   "Carrier_17_SpareSafetyInput(2_4)" AT %I1214.4 : Bool;   // SPARE SAFETY INPUT
   "Carrier_17_SpareSafetyInput(2_5)" AT %I1214.5 : Bool;   // SPARE SAFETY INPUT
   "Carrier_17_SpareSafetyInput(2_6)" AT %I1214.6 : Bool;   // SPARE SAFETY INPUT
   "Carrier_17_SpareSafetyInput(2_7)" AT %I1214.7 : Bool;   // SPARE SAFETY INPUT
   "Carrier_17_Slot3_SafetyOutput" AT %IW1215 : Word;   // SLOT 3 SAFETY OUTPUT WORD
   "Carrier_17_Crash_Detect_OK" AT %I1215.0 : Bool;   // CARRIER CRASH DETECT
   "Carrier_17_SpareSafetyOutput(3_1)" AT %I1215.1 : Bool;   // SPARE SAFETY OUTPUT
   "Carrier_17_SpareSafetyOutput(3_2)" AT %I1215.2 : Bool;   // SPARE SAFETY OUTPUT
   "Carrier_17_SpareSafetyOutput(3_3)" AT %I1215.3 : Bool;   // SPARE SAFETY OUTPUT
   "Carrier_17_SpareSafetyOutput(3_4)" AT %I1215.4 : Bool;   // SPARE SAFETY OUTPUT
   "Carrier_17_SpareSafetyOutput(3_5)" AT %I1215.5 : Bool;   // SPARE SAFETY OUTPUT
   "Carrier_17_SpareSafetyOutput(3_6)" AT %I1215.6 : Bool;   // SPARE SAFETY OUTPUT
   "Carrier_17_SpareSafetyOutput(3_7)" AT %I1215.7 : Bool;   // SPARE SAFETY OUTPUT
   "Carrier_17_Slot4_Input" AT %IW1216 : Word;   // SLOT 4 INPUT WORD
   "Carrier_17_480VPowerOn_MDCB1" AT %I1216.0 : Bool;   // 480 VAC POWER ON MDCB 1
   "Carrier_17_SpareInput(4_1)" AT %I1216.1 : Bool;   // SPARE INPUT
   "Carrier_17_SpareInput(4_2)" AT %I1216.2 : Bool;   // SPARE INPUT
   "Carrier_17_SitopSelectStatus" AT %I1216.3 : Bool;   // SITOP SELECT STATUS
   "Carrier_17_DCsupplyOnPSCB2" AT %I1216.4 : Bool;   // DC SUPPLY ON PSCB 2
   "Carrier_17_SpareInput(4_5)" AT %I1216.5 : Bool;   // SPARE INPUT
   "Carrier_17_SpareInput(4_6)" AT %I1216.6 : Bool;   // SPARE INPUT
   "Carrier_17_SpareInput(4_7)" AT %I1216.7 : Bool;   // SPARE INPUT
   "Carrier_17_PB1_ProdHoldLH" AT %I1217.0 : Bool;   // PB 1 PRODUCTION HOLD LH
   "Carrier_17_PB2_ResetLH" AT %I1217.1 : Bool;   // PB 2 RESET LH
   "Carrier_17_PB3_ProdHoldRH" AT %I1217.2 : Bool;   // PB 3 PRODUCTION HOLD RH
   "Carrier_17_PB4_ResetRH" AT %I1217.3 : Bool;   // PB 4 RESET RH
   "Carrier_17_SpareInput(4_14)" AT %I1217.4 : Bool;   // SPARE INPUT
   "Carrier_17_SpareInput(4_15)" AT %I1217.5 : Bool;   // SPARE INPUT
   "Carrier_17_SpareInput(4_16)" AT %I1217.6 : Bool;   // SPARE INPUT
   "Carrier_17_SpareInput(4_17)" AT %I1217.7 : Bool;   // SPARE INPUT
   "Carrier_17_Slot5_Output" AT %IW1218 : Word;   // SLOT 5 OUTPUT WORD
   "Carrier_17_IRD400_HMI_24VDC_ENABLE" AT %I1218.0 : Bool;   // IRD 400 PANEL HMI 24V DC POWER
   "Carrier_17_FaultLight_LH" AT %I1218.1 : Bool;   // FAULT LIGHT LH
   "Carrier_17_RunLight_LH" AT %I1218.2 : Bool;   // RUN LIGHT LH
   "Carrier_17_FaultLight_RH" AT %I1218.3 : Bool;   // FAULT LIGHT RH
   "Carrier_17_RunLight_RH" AT %I1218.4 : Bool;   // RUN LIGHT RH
   "Carrier_17_SpareOutput(5_5)" AT %I1218.5 : Bool;   // SPARE OUTPUT
   "Carrier_17_SpareOutput(5_6)" AT %I1218.6 : Bool;   // SPARE OUTPUT
   "Carrier_17_SpareOutput(5_7)" AT %I1218.7 : Bool;   // SPARE OUTPUT
   "Carrier_17_ActualSpeed" AT %IW1220 : Word;   // ACTUAL SPEED
   "Carrier_17_CarrierDriveAlarm" AT %IW1222 : Word;   // CARRIER DRIVE ALARM
   "Carrier_17_CarrierDriveWarning" AT %IW1224 : Word;   // CARRIER DRIVE WARNING
   "Carrier_18_Status" AT %IW1250 : Word;   // CARRIER STATUS WORD
   "Carrier_18_Status.0" AT %I1250.0 : Bool;   // HEARTBEAT
   "Carrier_18_Status.1" AT %I1250.1 : Bool;   // MANUAL
   "Carrier_18_Status.2" AT %I1250.2 : Bool;   // IN_AUTO
   "Carrier_18_Status.3" AT %I1250.3 : Bool;   // POSITIONING_COMPLETE
   "Carrier_18_Status.4" AT %I1250.4 : Bool;   // PRODUCTION HOLD
   "Carrier_18_Status.5" AT %I1250.5 : Bool;   // CARRIER MOVING FORWARD
   "Carrier_18_Status.6" AT %I1250.6 : Bool;   // CARRIER MOVING REVERSE
   "Carrier_18_Status.7" AT %I1250.7 : Bool;   // CARRIER FAULT
   "Carrier_18_Status.8" AT %I1251.0 : Bool;   // CRASH DETECT TRIPPED
   "Carrier_18_Status.9" AT %I1251.1 : Bool;
   "Carrier_18_Status.10" AT %I1251.2 : Bool;
   "Carrier_18_Status.11" AT %I1251.3 : Bool;
   "Carrier_18_Status.12" AT %I1251.4 : Bool;
   "Carrier_18_Status.13" AT %I1251.5 : Bool;
   "Carrier_18_Status.14" AT %I1251.6 : Bool;
   "Carrier_18_Status.15" AT %I1251.7 : Bool;
   "Carrier_18_SDCFaultCode" AT %IW1252 : Word;   // SDC FAULT CODE
   "Carrier_18_CarrierPosition" AT %ID1254 : DWord;   // CARRIER POSITION
   "Carrier_18_CarrierNumber" AT %IW1258 : Word;   // CARRIER NUMBER
   "Carrier_18_G120DControlWord" AT %IW1260 : Word;   // G120D_STW1_CONTROL
   "Carrier_18_G120DControlWord.0" AT %I1260.0 : Bool;   // Bit_00_ON
   "Carrier_18_G120DControlWord.1" AT %I1260.1 : Bool;   // Bit_01_AUS2_INH
   "Carrier_18_G120DControlWord.2" AT %I1260.2 : Bool;   // Bit_02_AUS3_STOP
   "Carrier_18_G120DControlWord.3" AT %I1260.3 : Bool;   // Bit_03_EN
   "Carrier_18_G120DControlWord.4" AT %I1260.4 : Bool;   // Bit_04_EN_RAMP
   "Carrier_18_G120DControlWord.5" AT %I1260.5 : Bool;   // Bit_05_START_RAMP
   "Carrier_18_G120DControlWord.6" AT %I1260.6 : Bool;   // Bit_06_SETPOINT
   "Carrier_18_G120DControlWord.7" AT %I1260.7 : Bool;   // Bit_07_RESET
   "Carrier_18_G120DControlWord.8" AT %I1261.0 : Bool;   // Bit_08_JOG_R
   "Carrier_18_G120DControlWord.9" AT %I1261.1 : Bool;   // Bit_09_JOG_L
   "Carrier_18_G120DControlWord.10" AT %I1261.2 : Bool;   // Bit_10_CONTR_PLC
   "Carrier_18_G120DControlWord.11" AT %I1261.3 : Bool;   // Bit_11_REVERSE
   "Carrier_18_G120DControlWord.12" AT %I1261.4 : Bool;   // Bit_12_BRAKE_RELEASE
   "Carrier_18_G120DControlWord.13" AT %I1261.5 : Bool;   // Bit_13_DDS
   "Carrier_18_G120DControlWord.14" AT %I1261.6 : Bool;   // Bit_14_DO0
   "Carrier_18_G120DControlWord.15" AT %I1261.7 : Bool;   // Bit_15_DO1
   "Carrier_18_G120DStatusWord" AT %IW1262 : Word;   // G120D_ZSW1_STATUS
   "Carrier_18_G120DStatusWord.0" AT %I1262.0 : Bool;   // Bit_00_READY_RUN
   "Carrier_18_G120DStatusWord.1" AT %I1262.1 : Bool;   // Bit_01_READY_ON
   "Carrier_18_G120DStatusWord.2" AT %I1262.2 : Bool;   // Bit_02_ENABLE
   "Carrier_18_G120DStatusWord.3" AT %I1262.3 : Bool;   // Bit_03_FAULT
   "Carrier_18_G120DStatusWord.4" AT %I1262.4 : Bool;   // Bit_04_OFF2
   "Carrier_18_G120DStatusWord.5" AT %I1262.5 : Bool;   // Bit_05_OFF3
   "Carrier_18_G120DStatusWord.6" AT %I1262.6 : Bool;   // Bit_06_LOCK_OUT
   "Carrier_18_G120DStatusWord.7" AT %I1262.7 : Bool;   // Bit_07_WARN
   "Carrier_18_G120DStatusWord.8" AT %I1263.0 : Bool;   // Bit_08_NO_DEVIATION
   "Carrier_18_G120DStatusWord.9" AT %I1263.1 : Bool;   // Bit_09_CONTR_PLC
   "Carrier_18_G120DStatusWord.10" AT %I1263.2 : Bool;   // Bit_10_F_MAX
   "Carrier_18_G120DStatusWord.11" AT %I1263.3 : Bool;   // Bit_11_LIMIT_REACHED
   "Carrier_18_G120DStatusWord.12" AT %I1263.4 : Bool;   // Bit_12_BRAKE_OPEN
   "Carrier_18_G120DStatusWord.13" AT %I1263.5 : Bool;   // Bit_13_NO_OVERTEMP
   "Carrier_18_G120DStatusWord.14" AT %I1263.6 : Bool;   // Bit_14_CW_CCW
   "Carrier_18_G120DStatusWord.15" AT %I1263.7 : Bool;   // Bit_15_OVERL
   "Carrier_18_Slot2_Input" AT %IW1264 : Word;   // SLOT 2 INPUT WORD
   "Carrier_18_CrashDetectSW" AT %I1264.0 : Bool;   // CRASH DETECT SW
   "Carrier_18_SpareSafetyInput(2_1)" AT %I1264.1 : Bool;   // SPARE SAFETY INPUT
   "Carrier_18_SpareSafetyInput(2_2)" AT %I1264.2 : Bool;   // SPARE SAFETY INPUT
   "Carrier_18_SpareSafetyInput(2_3)" AT %I1264.3 : Bool;   // SPARE SAFETY INPUT
   "Carrier_18_SpareSafetyInput(2_4)" AT %I1264.4 : Bool;   // SPARE SAFETY INPUT
   "Carrier_18_SpareSafetyInput(2_5)" AT %I1264.5 : Bool;   // SPARE SAFETY INPUT
   "Carrier_18_SpareSafetyInput(2_6)" AT %I1264.6 : Bool;   // SPARE SAFETY INPUT
   "Carrier_18_SpareSafetyInput(2_7)" AT %I1264.7 : Bool;   // SPARE SAFETY INPUT
   "Carrier_18_Slot3_SafetyOutput" AT %IW1265 : Word;   // SLOT 3 SAFETY OUTPUT WORD
   "Carrier_18_Crash_Detect_OK" AT %I1265.0 : Bool;   // CARRIER CRASH DETECT
   "Carrier_18_SpareSafetyOutput(3_1)" AT %I1265.1 : Bool;   // SPARE SAFETY OUTPUT
   "Carrier_18_SpareSafetyOutput(3_2)" AT %I1265.2 : Bool;   // SPARE SAFETY OUTPUT
   "Carrier_18_SpareSafetyOutput(3_3)" AT %I1265.3 : Bool;   // SPARE SAFETY OUTPUT
   "Carrier_18_SpareSafetyOutput(3_4)" AT %I1265.4 : Bool;   // SPARE SAFETY OUTPUT
   "Carrier_18_SpareSafetyOutput(3_5)" AT %I1265.5 : Bool;   // SPARE SAFETY OUTPUT
   "Carrier_18_SpareSafetyOutput(3_6)" AT %I1265.6 : Bool;   // SPARE SAFETY OUTPUT
   "Carrier_18_SpareSafetyOutput(3_7)" AT %I1265.7 : Bool;   // SPARE SAFETY OUTPUT
   "Carrier_18_Slot4_Input" AT %IW1266 : Word;   // SLOT 4 INPUT WORD
   "Carrier_18_480VPowerOn_MDCB1" AT %I1266.0 : Bool;   // 480 VAC POWER ON MDCB 1
   "Carrier_18_SpareInput(4_1)" AT %I1266.1 : Bool;   // SPARE INPUT
   "Carrier_18_SpareInput(4_2)" AT %I1266.2 : Bool;   // SPARE INPUT
   "Carrier_18_SitopSelectStatus" AT %I1266.3 : Bool;   // SITOP SELECT STATUS
   "Carrier_18_DCsupplyOnPSCB2" AT %I1266.4 : Bool;   // DC SUPPLY ON PSCB 2
   "Carrier_18_SpareInput(4_5)" AT %I1266.5 : Bool;   // SPARE INPUT
   "Carrier_18_SpareInput(4_6)" AT %I1266.6 : Bool;   // SPARE INPUT
   "Carrier_18_SpareInput(4_7)" AT %I1266.7 : Bool;   // SPARE INPUT
   "Carrier_18_PB1_ProdHoldLH" AT %I1267.0 : Bool;   // PB 1 PRODUCTION HOLD LH
   "Carrier_18_PB2_ResetLH" AT %I1267.1 : Bool;   // PB 2 RESET LH
   "Carrier_18_PB3_ProdHoldRH" AT %I1267.2 : Bool;   // PB 3 PRODUCTION HOLD RH
   "Carrier_18_PB4_ResetRH" AT %I1267.3 : Bool;   // PB 4 RESET RH
   "Carrier_18_SpareInput(4_14)" AT %I1267.4 : Bool;   // SPARE INPUT
   "Carrier_18_SpareInput(4_15)" AT %I1267.5 : Bool;   // SPARE INPUT
   "Carrier_18_SpareInput(4_16)" AT %I1267.6 : Bool;   // SPARE INPUT
   "Carrier_18_SpareInput(4_17)" AT %I1267.7 : Bool;   // SPARE INPUT
   "Carrier_18_Slot5_Output" AT %IW1268 : Word;   // SLOT 5 OUTPUT WORD
   "Carrier_18_IRD400_HMI_24VDC_ENABLE" AT %I1268.0 : Bool;   // IRD 400 PANEL HMI 24V DC POWER
   "Carrier_18_FaultLight_LH" AT %I1268.1 : Bool;   // FAULT LIGHT LH
   "Carrier_18_RunLight_LH" AT %I1268.2 : Bool;   // RUN LIGHT LH
   "Carrier_18_FaultLight_RH" AT %I1268.3 : Bool;   // FAULT LIGHT RH
   "Carrier_18_RunLight_RH" AT %I1268.4 : Bool;   // RUN LIGHT RH
   "Carrier_18_SpareOutput(5_5)" AT %I1268.5 : Bool;   // SPARE OUTPUT
   "Carrier_18_SpareOutput(5_6)" AT %I1268.6 : Bool;   // SPARE OUTPUT
   "Carrier_18_SpareOutput(5_7)" AT %I1268.7 : Bool;   // SPARE OUTPUT
   "Carrier_18_ActualSpeed" AT %IW1270 : Word;   // ACTUAL SPEED
   "Carrier_18_CarrierDriveAlarm" AT %IW1272 : Word;   // CARRIER DRIVE ALARM
   "Carrier_18_CarrierDriveWarning" AT %IW1274 : Word;   // CARRIER DRIVE WARNING
   "Carrier_19_Status" AT %IW1300 : Word;   // CARRIER STATUS WORD
   "Carrier_19_Status.0" AT %I1300.0 : Bool;   // HEARTBEAT
   "Carrier_19_Status.1" AT %I1300.1 : Bool;   // MANUAL
   "Carrier_19_Status.2" AT %I1300.2 : Bool;   // IN_AUTO
   "Carrier_19_Status.3" AT %I1300.3 : Bool;   // POSITIONING_COMPLETE
   "Carrier_19_Status.4" AT %I1300.4 : Bool;   // PRODUCTION HOLD
   "Carrier_19_Status.5" AT %I1300.5 : Bool;   // CARRIER MOVING FORWARD
   "Carrier_19_Status.6" AT %I1300.6 : Bool;   // CARRIER MOVING REVERSE
   "Carrier_19_Status.7" AT %I1300.7 : Bool;   // CARRIER FAULT
   "Carrier_19_Status.8" AT %I1301.0 : Bool;   // CRASH DETECT TRIPPED
   "Carrier_19_Status.9" AT %I1301.1 : Bool;
   "Carrier_19_Status.10" AT %I1301.2 : Bool;
   "Carrier_19_Status.11" AT %I1301.3 : Bool;
   "Carrier_19_Status.12" AT %I1301.4 : Bool;
   "Carrier_19_Status.13" AT %I1301.5 : Bool;
   "Carrier_19_Status.14" AT %I1301.6 : Bool;
   "Carrier_19_Status.15" AT %I1301.7 : Bool;
   "Carrier_19_SDCFaultCode" AT %IW1302 : Word;   // SDC FAULT CODE
   "Carrier_19_CarrierPosition" AT %ID1304 : DWord;   // CARRIER POSITION
   "Carrier_19_CarrierNumber" AT %IW1308 : Word;   // CARRIER NUMBER
   "Carrier_19_G120DControlWord" AT %IW1310 : Word;   // G120D_STW1_CONTROL
   "Carrier_19_G120DControlWord.0" AT %I1310.0 : Bool;   // Bit_00_ON
   "Carrier_19_G120DControlWord.1" AT %I1310.1 : Bool;   // Bit_01_AUS2_INH
   "Carrier_19_G120DControlWord.2" AT %I1310.2 : Bool;   // Bit_02_AUS3_STOP
   "Carrier_19_G120DControlWord.3" AT %I1310.3 : Bool;   // Bit_03_EN
   "Carrier_19_G120DControlWord.4" AT %I1310.4 : Bool;   // Bit_04_EN_RAMP
   "Carrier_19_G120DControlWord.5" AT %I1310.5 : Bool;   // Bit_05_START_RAMP
   "Carrier_19_G120DControlWord.6" AT %I1310.6 : Bool;   // Bit_06_SETPOINT
   "Carrier_19_G120DControlWord.7" AT %I1310.7 : Bool;   // Bit_07_RESET
   "Carrier_19_G120DControlWord.8" AT %I1311.0 : Bool;   // Bit_08_JOG_R
   "Carrier_19_G120DControlWord.9" AT %I1311.1 : Bool;   // Bit_09_JOG_L
   "Carrier_19_G120DControlWord.10" AT %I1311.2 : Bool;   // Bit_10_CONTR_PLC
   "Carrier_19_G120DControlWord.11" AT %I1311.3 : Bool;   // Bit_11_REVERSE
   "Carrier_19_G120DControlWord.12" AT %I1311.4 : Bool;   // Bit_12_BRAKE_RELEASE
   "Carrier_19_G120DControlWord.13" AT %I1311.5 : Bool;   // Bit_13_DDS
   "Carrier_19_G120DControlWord.14" AT %I1311.6 : Bool;   // Bit_14_DO0
   "Carrier_19_G120DControlWord.15" AT %I1311.7 : Bool;   // Bit_15_DO1
   "Carrier_19_G120DStatusWord" AT %IW1312 : Word;   // G120D_ZSW1_STATUS
   "Carrier_19_G120DStatusWord.0" AT %I1312.0 : Bool;   // Bit_00_READY_RUN
   "Carrier_19_G120DStatusWord.1" AT %I1312.1 : Bool;   // Bit_01_READY_ON
   "Carrier_19_G120DStatusWord.2" AT %I1312.2 : Bool;   // Bit_02_ENABLE
   "Carrier_19_G120DStatusWord.3" AT %I1312.3 : Bool;   // Bit_03_FAULT
   "Carrier_19_G120DStatusWord.4" AT %I1312.4 : Bool;   // Bit_04_OFF2
   "Carrier_19_G120DStatusWord.5" AT %I1312.5 : Bool;   // Bit_05_OFF3
   "Carrier_19_G120DStatusWord.6" AT %I1312.6 : Bool;   // Bit_06_LOCK_OUT
   "Carrier_19_G120DStatusWord.7" AT %I1312.7 : Bool;   // Bit_07_WARN
   "Carrier_19_G120DStatusWord.8" AT %I1313.0 : Bool;   // Bit_08_NO_DEVIATION
   "Carrier_19_G120DStatusWord.9" AT %I1313.1 : Bool;   // Bit_09_CONTR_PLC
   "Carrier_19_G120DStatusWord.10" AT %I1313.2 : Bool;   // Bit_10_F_MAX
   "Carrier_19_G120DStatusWord.11" AT %I1313.3 : Bool;   // Bit_11_LIMIT_REACHED
   "Carrier_19_G120DStatusWord.12" AT %I1313.4 : Bool;   // Bit_12_BRAKE_OPEN
   "Carrier_19_G120DStatusWord.13" AT %I1313.5 : Bool;   // Bit_13_NO_OVERTEMP
   "Carrier_19_G120DStatusWord.14" AT %I1313.6 : Bool;   // Bit_14_CW_CCW
   "Carrier_19_G120DStatusWord.15" AT %I1313.7 : Bool;   // Bit_15_OVERL
   "Carrier_19_Slot2_Input" AT %IW1314 : Word;   // SLOT 2 INPUT WORD
   "Carrier_19_CrashDetectSW" AT %I1314.0 : Bool;   // CRASH DETECT SW
   "Carrier_19_SpareSafetyInput(2_1)" AT %I1314.1 : Bool;   // SPARE SAFETY INPUT
   "Carrier_19_SpareSafetyInput(2_2)" AT %I1314.2 : Bool;   // SPARE SAFETY INPUT
   "Carrier_19_SpareSafetyInput(2_3)" AT %I1314.3 : Bool;   // SPARE SAFETY INPUT
   "Carrier_19_SpareSafetyInput(2_4)" AT %I1314.4 : Bool;   // SPARE SAFETY INPUT
   "Carrier_19_SpareSafetyInput(2_5)" AT %I1314.5 : Bool;   // SPARE SAFETY INPUT
   "Carrier_19_SpareSafetyInput(2_6)" AT %I1314.6 : Bool;   // SPARE SAFETY INPUT
   "Carrier_19_SpareSafetyInput(2_7)" AT %I1314.7 : Bool;   // SPARE SAFETY INPUT
   "Carrier_19_Slot3_SafetyOutput" AT %IW1315 : Word;   // SLOT 3 SAFETY OUTPUT WORD
   "Carrier_19_Crash_Detect_OK" AT %I1315.0 : Bool;   // CARRIER CRASH DETECT
   "Carrier_19_SpareSafetyOutput(3_1)" AT %I1315.1 : Bool;   // SPARE SAFETY OUTPUT
   "Carrier_19_SpareSafetyOutput(3_2)" AT %I1315.2 : Bool;   // SPARE SAFETY OUTPUT
   "Carrier_19_SpareSafetyOutput(3_3)" AT %I1315.3 : Bool;   // SPARE SAFETY OUTPUT
   "Carrier_19_SpareSafetyOutput(3_4)" AT %I1315.4 : Bool;   // SPARE SAFETY OUTPUT
   "Carrier_19_SpareSafetyOutput(3_5)" AT %I1315.5 : Bool;   // SPARE SAFETY OUTPUT
   "Carrier_19_SpareSafetyOutput(3_6)" AT %I1315.6 : Bool;   // SPARE SAFETY OUTPUT
   "Carrier_19_SpareSafetyOutput(3_7)" AT %I1315.7 : Bool;   // SPARE SAFETY OUTPUT
   "Carrier_19_Slot4_Input" AT %IW1316 : Word;   // SLOT 4 INPUT WORD
   "Carrier_19_480VPowerOn_MDCB1" AT %I1316.0 : Bool;   // 480 VAC POWER ON MDCB 1
   "Carrier_19_SpareInput(4_1)" AT %I1316.1 : Bool;   // SPARE INPUT
   "Carrier_19_SpareInput(4_2)" AT %I1316.2 : Bool;   // SPARE INPUT
   "Carrier_19_SitopSelectStatus" AT %I1316.3 : Bool;   // SITOP SELECT STATUS
   "Carrier_19_DCsupplyOnPSCB2" AT %I1316.4 : Bool;   // DC SUPPLY ON PSCB 2
   "Carrier_19_SpareInput(4_5)" AT %I1316.5 : Bool;   // SPARE INPUT
   "Carrier_19_SpareInput(4_6)" AT %I1316.6 : Bool;   // SPARE INPUT
   "Carrier_19_SpareInput(4_7)" AT %I1316.7 : Bool;   // SPARE INPUT
   "Carrier_19_PB1_ProdHoldLH" AT %I1317.0 : Bool;   // PB 1 PRODUCTION HOLD LH
   "Carrier_19_PB2_ResetLH" AT %I1317.1 : Bool;   // PB 2 RESET LH
   "Carrier_19_PB3_ProdHoldRH" AT %I1317.2 : Bool;   // PB 3 PRODUCTION HOLD RH
   "Carrier_19_PB4_ResetRH" AT %I1317.3 : Bool;   // PB 4 RESET RH
   "Carrier_19_SpareInput(4_14)" AT %I1317.4 : Bool;   // SPARE INPUT
   "Carrier_19_SpareInput(4_15)" AT %I1317.5 : Bool;   // SPARE INPUT
   "Carrier_19_SpareInput(4_16)" AT %I1317.6 : Bool;   // SPARE INPUT
   "Carrier_19_SpareInput(4_17)" AT %I1317.7 : Bool;   // SPARE INPUT
   "Carrier_19_Slot5_Output" AT %IW1318 : Word;   // SLOT 5 OUTPUT WORD
   "Carrier_19_IRD400_HMI_24VDC_ENABLE" AT %I1318.0 : Bool;   // IRD 400 PANEL HMI 24V DC POWER
   "Carrier_19_FaultLight_LH" AT %I1318.1 : Bool;   // FAULT LIGHT LH
   "Carrier_19_RunLight_LH" AT %I1318.2 : Bool;   // RUN LIGHT LH
   "Carrier_19_FaultLight_RH" AT %I1318.3 : Bool;   // FAULT LIGHT RH
   "Carrier_19_RunLight_RH" AT %I1318.4 : Bool;   // RUN LIGHT RH
   "Carrier_19_SpareOutput(5_5)" AT %I1318.5 : Bool;   // SPARE OUTPUT
   "Carrier_19_SpareOutput(5_6)" AT %I1318.6 : Bool;   // SPARE OUTPUT
   "Carrier_19_SpareOutput(5_7)" AT %I1318.7 : Bool;   // SPARE OUTPUT
   "Carrier_19_ActualSpeed" AT %IW1320 : Word;   // ACTUAL SPEED
   "Carrier_19_CarrierDriveAlarm" AT %IW1322 : Word;   // CARRIER DRIVE ALARM
   "Carrier_19_CarrierDriveWarning" AT %IW1324 : Word;   // CARRIER DRIVE WARNING
   "Carrier_20_Status" AT %IW1350 : Word;   // CARRIER STATUS WORD
   "Carrier_20_Status.0" AT %I1350.0 : Bool;   // HEARTBEAT
   "Carrier_20_Status.1" AT %I1350.1 : Bool;   // MANUAL
   "Carrier_20_Status.2" AT %I1350.2 : Bool;   // IN_AUTO
   "Carrier_20_Status.3" AT %I1350.3 : Bool;   // POSITIONING_COMPLETE
   "Carrier_20_Status.4" AT %I1350.4 : Bool;   // PRODUCTION HOLD
   "Carrier_20_Status.5" AT %I1350.5 : Bool;   // CARRIER MOVING FORWARD
   "Carrier_20_Status.6" AT %I1350.6 : Bool;   // CARRIER MOVING REVERSE
   "Carrier_20_Status.7" AT %I1350.7 : Bool;   // CARRIER FAULT
   "Carrier_20_Status.8" AT %I1351.0 : Bool;   // CRASH DETECT TRIPPED
   "Carrier_20_Status.9" AT %I1351.1 : Bool;
   "Carrier_20_Status.10" AT %I1351.2 : Bool;
   "Carrier_20_Status.11" AT %I1351.3 : Bool;
   "Carrier_20_Status.12" AT %I1351.4 : Bool;
   "Carrier_20_Status.13" AT %I1351.5 : Bool;
   "Carrier_20_Status.14" AT %I1351.6 : Bool;
   "Carrier_20_Status.15" AT %I1351.7 : Bool;
   "Carrier_20_SDCFaultCode" AT %IW1352 : Word;   // SDC FAULT CODE
   "Carrier_20_CarrierPosition" AT %ID1354 : DWord;   // CARRIER POSITION
   "Carrier_20_CarrierNumber" AT %IW1358 : Word;   // CARRIER NUMBER
   "Carrier_20_G120DControlWord" AT %IW1360 : Word;   // G120D_STW1_CONTROL
   "Carrier_20_G120DControlWord.0" AT %I1360.0 : Bool;   // Bit_00_ON
   "Carrier_20_G120DControlWord.1" AT %I1360.1 : Bool;   // Bit_01_AUS2_INH
   "Carrier_20_G120DControlWord.2" AT %I1360.2 : Bool;   // Bit_02_AUS3_STOP
   "Carrier_20_G120DControlWord.3" AT %I1360.3 : Bool;   // Bit_03_EN
   "Carrier_20_G120DControlWord.4" AT %I1360.4 : Bool;   // Bit_04_EN_RAMP
   "Carrier_20_G120DControlWord.5" AT %I1360.5 : Bool;   // Bit_05_START_RAMP
   "Carrier_20_G120DControlWord.6" AT %I1360.6 : Bool;   // Bit_06_SETPOINT
   "Carrier_20_G120DControlWord.7" AT %I1360.7 : Bool;   // Bit_07_RESET
   "Carrier_20_G120DControlWord.8" AT %I1361.0 : Bool;   // Bit_08_JOG_R
   "Carrier_20_G120DControlWord.9" AT %I1361.1 : Bool;   // Bit_09_JOG_L
   "Carrier_20_G120DControlWord.10" AT %I1361.2 : Bool;   // Bit_10_CONTR_PLC
   "Carrier_20_G120DControlWord.11" AT %I1361.3 : Bool;   // Bit_11_REVERSE
   "Carrier_20_G120DControlWord.12" AT %I1361.4 : Bool;   // Bit_12_BRAKE_RELEASE
   "Carrier_20_G120DControlWord.13" AT %I1361.5 : Bool;   // Bit_13_DDS
   "Carrier_20_G120DControlWord.14" AT %I1361.6 : Bool;   // Bit_14_DO0
   "Carrier_20_G120DControlWord.15" AT %I1361.7 : Bool;   // Bit_15_DO1
   "Carrier_20_G120DStatusWord" AT %IW1362 : Word;   // G120D_ZSW1_STATUS
   "Carrier_20_G120DStatusWord.0" AT %I1362.0 : Bool;   // Bit_00_READY_RUN
   "Carrier_20_G120DStatusWord.1" AT %I1362.1 : Bool;   // Bit_01_READY_ON
   "Carrier_20_G120DStatusWord.2" AT %I1362.2 : Bool;   // Bit_02_ENABLE
   "Carrier_20_G120DStatusWord.3" AT %I1362.3 : Bool;   // Bit_03_FAULT
   "Carrier_20_G120DStatusWord.4" AT %I1362.4 : Bool;   // Bit_04_OFF2
   "Carrier_20_G120DStatusWord.5" AT %I1362.5 : Bool;   // Bit_05_OFF3
   "Carrier_20_G120DStatusWord.6" AT %I1362.6 : Bool;   // Bit_06_LOCK_OUT
   "Carrier_20_G120DStatusWord.7" AT %I1362.7 : Bool;   // Bit_07_WARN
   "Carrier_20_G120DStatusWord.8" AT %I1363.0 : Bool;   // Bit_08_NO_DEVIATION
   "Carrier_20_G120DStatusWord.9" AT %I1363.1 : Bool;   // Bit_09_CONTR_PLC
   "Carrier_20_G120DStatusWord.10" AT %I1363.2 : Bool;   // Bit_10_F_MAX
   "Carrier_20_G120DStatusWord.11" AT %I1363.3 : Bool;   // Bit_11_LIMIT_REACHED
   "Carrier_20_G120DStatusWord.12" AT %I1363.4 : Bool;   // Bit_12_BRAKE_OPEN
   "Carrier_20_G120DStatusWord.13" AT %I1363.5 : Bool;   // Bit_13_NO_OVERTEMP
   "Carrier_20_G120DStatusWord.14" AT %I1363.6 : Bool;   // Bit_14_CW_CCW
   "Carrier_20_G120DStatusWord.15" AT %I1363.7 : Bool;   // Bit_15_OVERL
   "Carrier_20_Slot2_Input" AT %IW1364 : Word;   // SLOT 2 INPUT WORD
   "Carrier_20_CrashDetectSW" AT %I1364.0 : Bool;   // CRASH DETECT SW
   "Carrier_20_SpareSafetyInput(2_1)" AT %I1364.1 : Bool;   // SPARE SAFETY INPUT
   "Carrier_20_SpareSafetyInput(2_2)" AT %I1364.2 : Bool;   // SPARE SAFETY INPUT
   "Carrier_20_SpareSafetyInput(2_3)" AT %I1364.3 : Bool;   // SPARE SAFETY INPUT
   "Carrier_20_SpareSafetyInput(2_4)" AT %I1364.4 : Bool;   // SPARE SAFETY INPUT
   "Carrier_20_SpareSafetyInput(2_5)" AT %I1364.5 : Bool;   // SPARE SAFETY INPUT
   "Carrier_20_SpareSafetyInput(2_6)" AT %I1364.6 : Bool;   // SPARE SAFETY INPUT
   "Carrier_20_SpareSafetyInput(2_7)" AT %I1364.7 : Bool;   // SPARE SAFETY INPUT
   "Carrier_20_Slot3_SafetyOutput" AT %IW1365 : Word;   // SLOT 3 SAFETY OUTPUT WORD
   "Carrier_20_Crash_Detect_OK" AT %I1365.0 : Bool;   // CARRIER CRASH DETECT
   "Carrier_20_SpareSafetyOutput(3_1)" AT %I1365.1 : Bool;   // SPARE SAFETY OUTPUT
   "Carrier_20_SpareSafetyOutput(3_2)" AT %I1365.2 : Bool;   // SPARE SAFETY OUTPUT
   "Carrier_20_SpareSafetyOutput(3_3)" AT %I1365.3 : Bool;   // SPARE SAFETY OUTPUT
   "Carrier_20_SpareSafetyOutput(3_4)" AT %I1365.4 : Bool;   // SPARE SAFETY OUTPUT
   "Carrier_20_SpareSafetyOutput(3_5)" AT %I1365.5 : Bool;   // SPARE SAFETY OUTPUT
   "Carrier_20_SpareSafetyOutput(3_6)" AT %I1365.6 : Bool;   // SPARE SAFETY OUTPUT
   "Carrier_20_SpareSafetyOutput(3_7)" AT %I1365.7 : Bool;   // SPARE SAFETY OUTPUT
   "Carrier_20_Slot4_Input" AT %IW1366 : Word;   // SLOT 4 INPUT WORD
   "Carrier_20_480VPowerOn_MDCB1" AT %I1366.0 : Bool;   // 480 VAC POWER ON MDCB 1
   "Carrier_20_SpareInput(4_1)" AT %I1366.1 : Bool;   // SPARE INPUT
   "Carrier_20_SpareInput(4_2)" AT %I1366.2 : Bool;   // SPARE INPUT
   "Carrier_20_SitopSelectStatus" AT %I1366.3 : Bool;   // SITOP SELECT STATUS
   "Carrier_20_DCsupplyOnPSCB2" AT %I1366.4 : Bool;   // DC SUPPLY ON PSCB 2
   "Carrier_20_SpareInput(4_5)" AT %I1366.5 : Bool;   // SPARE INPUT
   "Carrier_20_SpareInput(4_6)" AT %I1366.6 : Bool;   // SPARE INPUT
   "Carrier_20_SpareInput(4_7)" AT %I1366.7 : Bool;   // SPARE INPUT
   "Carrier_20_PB1_ProdHoldLH" AT %I1367.0 : Bool;   // PB 1 PRODUCTION HOLD LH
   "Carrier_20_PB2_ResetLH" AT %I1367.1 : Bool;   // PB 2 RESET LH
   "Carrier_20_PB3_ProdHoldRH" AT %I1367.2 : Bool;   // PB 3 PRODUCTION HOLD RH
   "Carrier_20_PB4_ResetRH" AT %I1367.3 : Bool;   // PB 4 RESET RH
   "Carrier_20_SpareInput(4_14)" AT %I1367.4 : Bool;   // SPARE INPUT
   "Carrier_20_SpareInput(4_15)" AT %I1367.5 : Bool;   // SPARE INPUT
   "Carrier_20_SpareInput(4_16)" AT %I1367.6 : Bool;   // SPARE INPUT
   "Carrier_20_SpareInput(4_17)" AT %I1367.7 : Bool;   // SPARE INPUT
   "Carrier_20_Slot5_Output" AT %IW1368 : Word;   // SLOT 5 OUTPUT WORD
   "Carrier_20_IRD400_HMI_24VDC_ENABLE" AT %I1368.0 : Bool;   // IRD 400 PANEL HMI 24V DC POWER
   "Carrier_20_FaultLight_LH" AT %I1368.1 : Bool;   // FAULT LIGHT LH
   "Carrier_20_RunLight_LH" AT %I1368.2 : Bool;   // RUN LIGHT LH
   "Carrier_20_FaultLight_RH" AT %I1368.3 : Bool;   // FAULT LIGHT RH
   "Carrier_20_RunLight_RH" AT %I1368.4 : Bool;   // RUN LIGHT RH
   "Carrier_20_SpareOutput(5_5)" AT %I1368.5 : Bool;   // SPARE OUTPUT
   "Carrier_20_SpareOutput(5_6)" AT %I1368.6 : Bool;   // SPARE OUTPUT
   "Carrier_20_SpareOutput(5_7)" AT %I1368.7 : Bool;   // SPARE OUTPUT
   "Carrier_20_ActualSpeed" AT %IW1370 : Word;   // ACTUAL SPEED
   "Carrier_20_CarrierDriveAlarm" AT %IW1372 : Word;   // CARRIER DRIVE ALARM
   "Carrier_20_CarrierDriveWarning" AT %IW1374 : Word;   // CARRIER DRIVE WARNING
   "Carrier_21_Status" AT %IW1400 : Word;   // CARRIER STATUS WORD
   "Carrier_21_Status.0" AT %I1400.0 : Bool;   // HEARTBEAT
   "Carrier_21_Status.1" AT %I1400.1 : Bool;   // MANUAL
   "Carrier_21_Status.2" AT %I1400.2 : Bool;   // IN_AUTO
   "Carrier_21_Status.3" AT %I1400.3 : Bool;   // POSITIONING_COMPLETE
   "Carrier_21_Status.4" AT %I1400.4 : Bool;   // PRODUCTION HOLD
   "Carrier_21_Status.5" AT %I1400.5 : Bool;   // CARRIER MOVING FORWARD
   "Carrier_21_Status.6" AT %I1400.6 : Bool;   // CARRIER MOVING REVERSE
   "Carrier_21_Status.7" AT %I1400.7 : Bool;   // CARRIER FAULT
   "Carrier_21_Status.8" AT %I1401.0 : Bool;   // CRASH DETECT TRIPPED
   "Carrier_21_Status.9" AT %I1401.1 : Bool;
   "Carrier_21_Status.10" AT %I1401.2 : Bool;
   "Carrier_21_Status.11" AT %I1401.3 : Bool;
   "Carrier_21_Status.12" AT %I1401.4 : Bool;
   "Carrier_21_Status.13" AT %I1401.5 : Bool;
   "Carrier_21_Status.14" AT %I1401.6 : Bool;
   "Carrier_21_Status.15" AT %I1401.7 : Bool;
   "Carrier_21_SDCFaultCode" AT %IW1402 : Word;   // SDC FAULT CODE
   "Carrier_21_CarrierPosition" AT %ID1404 : DWord;   // CARRIER POSITION
   "Carrier_21_CarrierNumber" AT %IW1408 : Word;   // CARRIER NUMBER
   "Carrier_21_G120DControlWord" AT %IW1410 : Word;   // G120D_STW1_CONTROL
   "Carrier_21_G120DControlWord.0" AT %I1410.0 : Bool;   // Bit_00_ON
   "Carrier_21_G120DControlWord.1" AT %I1410.1 : Bool;   // Bit_01_AUS2_INH
   "Carrier_21_G120DControlWord.2" AT %I1410.2 : Bool;   // Bit_02_AUS3_STOP
   "Carrier_21_G120DControlWord.3" AT %I1410.3 : Bool;   // Bit_03_EN
   "Carrier_21_G120DControlWord.4" AT %I1410.4 : Bool;   // Bit_04_EN_RAMP
   "Carrier_21_G120DControlWord.5" AT %I1410.5 : Bool;   // Bit_05_START_RAMP
   "Carrier_21_G120DControlWord.6" AT %I1410.6 : Bool;   // Bit_06_SETPOINT
   "Carrier_21_G120DControlWord.7" AT %I1410.7 : Bool;   // Bit_07_RESET
   "Carrier_21_G120DControlWord.8" AT %I1411.0 : Bool;   // Bit_08_JOG_R
   "Carrier_21_G120DControlWord.9" AT %I1411.1 : Bool;   // Bit_09_JOG_L
   "Carrier_21_G120DControlWord.10" AT %I1411.2 : Bool;   // Bit_10_CONTR_PLC
   "Carrier_21_G120DControlWord.11" AT %I1411.3 : Bool;   // Bit_11_REVERSE
   "Carrier_21_G120DControlWord.12" AT %I1411.4 : Bool;   // Bit_12_BRAKE_RELEASE
   "Carrier_21_G120DControlWord.13" AT %I1411.5 : Bool;   // Bit_13_DDS
   "Carrier_21_G120DControlWord.14" AT %I1411.6 : Bool;   // Bit_14_DO0
   "Carrier_21_G120DControlWord.15" AT %I1411.7 : Bool;   // Bit_15_DO1
   "Carrier_21_G120DStatusWord" AT %IW1412 : Word;   // G120D_ZSW1_STATUS
   "Carrier_21_G120DStatusWord.0" AT %I1412.0 : Bool;   // Bit_00_READY_RUN
   "Carrier_21_G120DStatusWord.1" AT %I1412.1 : Bool;   // Bit_01_READY_ON
   "Carrier_21_G120DStatusWord.2" AT %I1412.2 : Bool;   // Bit_02_ENABLE
   "Carrier_21_G120DStatusWord.3" AT %I1412.3 : Bool;   // Bit_03_FAULT
   "Carrier_21_G120DStatusWord.4" AT %I1412.4 : Bool;   // Bit_04_OFF2
   "Carrier_21_G120DStatusWord.5" AT %I1412.5 : Bool;   // Bit_05_OFF3
   "Carrier_21_G120DStatusWord.6" AT %I1412.6 : Bool;   // Bit_06_LOCK_OUT
   "Carrier_21_G120DStatusWord.7" AT %I1412.7 : Bool;   // Bit_07_WARN
   "Carrier_21_G120DStatusWord.8" AT %I1413.0 : Bool;   // Bit_08_NO_DEVIATION
   "Carrier_21_G120DStatusWord.9" AT %I1413.1 : Bool;   // Bit_09_CONTR_PLC
   "Carrier_21_G120DStatusWord.10" AT %I1413.2 : Bool;   // Bit_10_F_MAX
   "Carrier_21_G120DStatusWord.11" AT %I1413.3 : Bool;   // Bit_11_LIMIT_REACHED
   "Carrier_21_G120DStatusWord.12" AT %I1413.4 : Bool;   // Bit_12_BRAKE_OPEN
   "Carrier_21_G120DStatusWord.13" AT %I1413.5 : Bool;   // Bit_13_NO_OVERTEMP
   "Carrier_21_G120DStatusWord.14" AT %I1413.6 : Bool;   // Bit_14_CW_CCW
   "Carrier_21_G120DStatusWord.15" AT %I1413.7 : Bool;   // Bit_15_OVERL
   "Carrier_21_Slot2_Input" AT %IW1414 : Word;   // SLOT 2 INPUT WORD
   "Carrier_21_CrashDetectSW" AT %I1414.0 : Bool;   // CRASH DETECT SW
   "Carrier_21_SpareSafetyInput(2_1)" AT %I1414.1 : Bool;   // SPARE SAFETY INPUT
   "Carrier_21_SpareSafetyInput(2_2)" AT %I1414.2 : Bool;   // SPARE SAFETY INPUT
   "Carrier_21_SpareSafetyInput(2_3)" AT %I1414.3 : Bool;   // SPARE SAFETY INPUT
   "Carrier_21_SpareSafetyInput(2_4)" AT %I1414.4 : Bool;   // SPARE SAFETY INPUT
   "Carrier_21_SpareSafetyInput(2_5)" AT %I1414.5 : Bool;   // SPARE SAFETY INPUT
   "Carrier_21_SpareSafetyInput(2_6)" AT %I1414.6 : Bool;   // SPARE SAFETY INPUT
   "Carrier_21_SpareSafetyInput(2_7)" AT %I1414.7 : Bool;   // SPARE SAFETY INPUT
   "Carrier_21_Slot3_SafetyOutput" AT %IW1415 : Word;   // SLOT 3 SAFETY OUTPUT WORD
   "Carrier_21_Crash_Detect_OK" AT %I1415.0 : Bool;   // CARRIER CRASH DETECT
   "Carrier_21_SpareSafetyOutput(3_1)" AT %I1415.1 : Bool;   // SPARE SAFETY OUTPUT
   "Carrier_21_SpareSafetyOutput(3_2)" AT %I1415.2 : Bool;   // SPARE SAFETY OUTPUT
   "Carrier_21_SpareSafetyOutput(3_3)" AT %I1415.3 : Bool;   // SPARE SAFETY OUTPUT
   "Carrier_21_SpareSafetyOutput(3_4)" AT %I1415.4 : Bool;   // SPARE SAFETY OUTPUT
   "Carrier_21_SpareSafetyOutput(3_5)" AT %I1415.5 : Bool;   // SPARE SAFETY OUTPUT
   "Carrier_21_SpareSafetyOutput(3_6)" AT %I1415.6 : Bool;   // SPARE SAFETY OUTPUT
   "Carrier_21_SpareSafetyOutput(3_7)" AT %I1415.7 : Bool;   // SPARE SAFETY OUTPUT
   "Carrier_21_Slot4_Input" AT %IW1416 : Word;   // SLOT 4 INPUT WORD
   "Carrier_21_480VPowerOn_MDCB1" AT %I1416.0 : Bool;   // 480 VAC POWER ON MDCB 1
   "Carrier_21_SpareInput(4_1)" AT %I1416.1 : Bool;   // SPARE INPUT
   "Carrier_21_SpareInput(4_2)" AT %I1416.2 : Bool;   // SPARE INPUT
   "Carrier_21_SitopSelectStatus" AT %I1416.3 : Bool;   // SITOP SELECT STATUS
   "Carrier_21_DCsupplyOnPSCB2" AT %I1416.4 : Bool;   // DC SUPPLY ON PSCB 2
   "Carrier_21_SpareInput(4_5)" AT %I1416.5 : Bool;   // SPARE INPUT
   "Carrier_21_SpareInput(4_6)" AT %I1416.6 : Bool;   // SPARE INPUT
   "Carrier_21_SpareInput(4_7)" AT %I1416.7 : Bool;   // SPARE INPUT
   "Carrier_21_PB1_ProdHoldLH" AT %I1417.0 : Bool;   // PB 1 PRODUCTION HOLD LH
   "Carrier_21_PB2_ResetLH" AT %I1417.1 : Bool;   // PB 2 RESET LH
   "Carrier_21_PB3_ProdHoldRH" AT %I1417.2 : Bool;   // PB 3 PRODUCTION HOLD RH
   "Carrier_21_PB4_ResetRH" AT %I1417.3 : Bool;   // PB 4 RESET RH
   "Carrier_21_SpareInput(4_14)" AT %I1417.4 : Bool;   // SPARE INPUT
   "Carrier_21_SpareInput(4_15)" AT %I1417.5 : Bool;   // SPARE INPUT
   "Carrier_21_SpareInput(4_16)" AT %I1417.6 : Bool;   // SPARE INPUT
   "Carrier_21_SpareInput(4_17)" AT %I1417.7 : Bool;   // SPARE INPUT
   "Carrier_21_Slot5_Output" AT %IW1418 : Word;   // SLOT 5 OUTPUT WORD
   "Carrier_21_IRD400_HMI_24VDC_ENABLE" AT %I1418.0 : Bool;   // IRD 400 PANEL HMI 24V DC POWER
   "Carrier_21_FaultLight_LH" AT %I1418.1 : Bool;   // FAULT LIGHT LH
   "Carrier_21_RunLight_LH" AT %I1418.2 : Bool;   // RUN LIGHT LH
   "Carrier_21_FaultLight_RH" AT %I1418.3 : Bool;   // FAULT LIGHT RH
   "Carrier_21_RunLight_RH" AT %I1418.4 : Bool;   // RUN LIGHT RH
   "Carrier_21_SpareOutput(5_5)" AT %I1418.5 : Bool;   // SPARE OUTPUT
   "Carrier_21_SpareOutput(5_6)" AT %I1418.6 : Bool;   // SPARE OUTPUT
   "Carrier_21_SpareOutput(5_7)" AT %I1418.7 : Bool;   // SPARE OUTPUT
   "Carrier_21_ActualSpeed" AT %IW1420 : Word;   // ACTUAL SPEED
   "Carrier_21_CarrierDriveAlarm" AT %IW1422 : Word;   // CARRIER DRIVE ALARM
   "Carrier_21_CarrierDriveWarning" AT %IW1424 : Word;   // CARRIER DRIVE WARNING
   "Carrier_22_Status" AT %IW1450 : Word;   // CARRIER STATUS WORD
   "Carrier_22_Status.0" AT %I1450.0 : Bool;   // HEARTBEAT
   "Carrier_22_Status.1" AT %I1450.1 : Bool;   // MANUAL
   "Carrier_22_Status.2" AT %I1450.2 : Bool;   // IN_AUTO
   "Carrier_22_Status.3" AT %I1450.3 : Bool;   // POSITIONING_COMPLETE
   "Carrier_22_Status.4" AT %I1450.4 : Bool;   // PRODUCTION HOLD
   "Carrier_22_Status.5" AT %I1450.5 : Bool;   // CARRIER MOVING FORWARD
   "Carrier_22_Status.6" AT %I1450.6 : Bool;   // CARRIER MOVING REVERSE
   "Carrier_22_Status.7" AT %I1450.7 : Bool;   // CARRIER FAULT
   "Carrier_22_Status.8" AT %I1451.0 : Bool;   // CRASH DETECT TRIPPED
   "Carrier_22_Status.9" AT %I1451.1 : Bool;
   "Carrier_22_Status.10" AT %I1451.2 : Bool;
   "Carrier_22_Status.11" AT %I1451.3 : Bool;
   "Carrier_22_Status.12" AT %I1451.4 : Bool;
   "Carrier_22_Status.13" AT %I1451.5 : Bool;
   "Carrier_22_Status.14" AT %I1451.6 : Bool;